// TIA Portal project "HEAT-1-CADIZ-V30" (V20) (continued)
VERSION : 0.1
// stored: InstanceOfName ToolChange
"ToolChange"
BEGIN
END_DATA_BLOCK

DATA_BLOCK "ToolChangeMarker_DB"   // DB40
{ S7_Optimized_Access := 'TRUE' }
VERSION : 0.1
// stored: InstanceOfName ToolChange
"ToolChange"
BEGIN
END_DATA_BLOCK

// folder: 30. Safety

DATA_BLOCK "InstMainSafety"   // DB1, F_DB
{ S7_Optimized_Access := 'TRUE' }
NAME : FUSI
VERSION : 0.1
// stored: InstanceOfName MainSafety
"MainSafety"
BEGIN
END_DATA_BLOCK

DATA_BLOCK "SafetyRobotDb"   // DB3, F_DB
{ S7_Optimized_Access := 'TRUE' }
VERSION : 0.1
BEGIN
END_DATA_BLOCK

DATA_BLOCK "EMERGENCIA_OPR_DB"   // DB41, F_DB
{ S7_Optimized_Access := 'TRUE' }
VERSION : 0.1
// stored: InstanceOfName EMERGENCIA_OPR
"EMERGENCIA_OPR"
BEGIN
END_DATA_BLOCK

DATA_BLOCK "EMERGENCIA_SETAS_DB"   // DB42, F_DB
{ S7_Optimized_Access := 'TRUE' }
VERSION : 0.1
// stored: InstanceOfName EMERGENCIA_SETAS
"EMERGENCIA_SETAS"
BEGIN
END_DATA_BLOCK

DATA_BLOCK "EMERGENCIAS_ANTENAS_DB"   // DB43, F_DB
{ S7_Optimized_Access := 'TRUE' }
VERSION : 0.1
// stored: InstanceOfName EMERGENCIAS_ANTENAS
"EMERGENCIAS_ANTENAS"
BEGIN
END_DATA_BLOCK

DATA_BLOCK "EMERGENCIA_GENERAL_DB"   // DB45, F_DB
{ S7_Optimized_Access := 'TRUE' }
VERSION : 0.1
// stored: InstanceOfName EMERGENCIA_GENERAL
"EMERGENCIA_GENERAL"
BEGIN
END_DATA_BLOCK

DATA_BLOCK "GESTION_BARRERAS_DB"   // DB46, F_DB
{ S7_Optimized_Access := 'TRUE' }
VERSION : 0.1
// stored: InstanceOfName GESTION_BARRERAS
"GESTION_BARRERAS"
BEGIN
END_DATA_BLOCK

// folder: 410. Festo cuba

DATA_BLOCK "HMI_CUBA_FESTO"   // DB12
{ S7_Optimized_Access := 'TRUE' }
VERSION : 0.1
   VAR
      HMI_Sensor_plato_giro_1 : Bool;
      HMI_Sensor_Plato_giro_2 : Bool;
      HMI_Sensor_plato_giro_3 : Bool;
      HMI_Sensor_ADN_bastidor_bloqueado_1 : Bool;
      HMI_Sensor_ADN_bastidor_desbloqueado_1 : Bool;
      HMI_Sensor_ADN_bastidor_bloqueado_2 : Bool;
      HMI_Sensor_ADN_bastidor_desbloqueado_2 : Bool;
      HMI_SENSOR_CRDSNU_BASTIDOR_BLOQUEADO_1 : Bool;
      HMI_SENSOR_CRDSNU_BASTIDOR_DESBLOQUEADO_1 : Bool;
      HMI_SENSOR_CRDSNU_BASTIDOR_BLOQUEADO_2 : Bool;
      HMI_SENSOR_CRDSNU_BASTIDOR_DESBLOQUEADO_2 : Bool;
      HMI_SENSOR_DSBG_BASTIDOR_ARRIBA_1 : Bool;
      HMI_SENSOR_DSBG_BASTIDOR_ABAJO_1 : Bool;
      HMI_SENSOR_DSBG_BASTIDOR_ARRIBA_2 : Bool;
      HMI_SENSOR_DSBG_BASTIDOR_ABAJO_2 : Bool;
      HMI_PULSADOR_SUBIR_1 : Bool;
      HMI_PULSADOR_BAJAR_1 : Bool;
      HMI_PULSADOR_SUBIR_2 : Bool;
      HMI_PULSADOR_BAJAR_2 : Bool;
      HMI_PULSADOR_BAJAR_3 : Bool;
      HMI_PULSADOR_BAJAR_4 : Bool;
      HMI_PULSADOR_BAJAR_5 : Bool;
      HMI_PULSADOR_BAJAR_6 : Bool;
      HMI_PULSADOR_BAJAR_7 : Bool;
      HMI_PULSADOR_BAJAR_8 : Bool;
      HMI_PULSADOR_BAJAR_9 : Bool;
      HMI_PULSADOR_BAJAR_10 : Bool;
      HMI_PULSADOR_BAJAR_11 : Bool;
      HMI_PULSADOR_BAJAR_12 : Bool;
      HMI_PULSADOR_BAJAR_13 : Bool;
      HMI_PULSADOR_BAJAR_14 : Bool;
      HMI_VALVULA_52_BIESTABLE_11 : Bool;
      HMI_VALVULA_52_BIESTABLE_12 : Bool;
      HMI_VALVULA_52_BIESTABLE_21 : Bool;
      HMI_VALVULA_52_BIESTABLE_22 : Bool;
      HMI_VÁLVULA_52_MONOESTABLE_1 : Bool;
      HMI_VÁLVULA_52_MONOESTABLE_2 : Bool;
      HMI_VÁLVULA_52_MONOESTABLE_3 : Bool;
      HMI_VÁLVULA_52_MONOESTABLE_4 : Bool;
      HMI_VÁLVULA_52_MONOESTABLE_5 : Bool;
      HMI_VÁLVULA_52_MONOESTABLE_6 : Bool;
      HMI_VÁLVULA_52_MONOESTABLE_7 : Bool;
      HMI_VÁLVULA_52_MONOESTABLE_8 : Bool;
      HMI_VÁLVULA_52_MONOESTABLE_9 : Bool;
      HMI_VÁLVULA_52_MONOESTABLE_10 : Bool;
      HMI_VÁLVULA_52_MONOESTABLE_11 : Bool;
      HMI_VÁLVULA_52_MONOESTABLE_12 : Bool;
      HMI_VÁLVULA_52_MONOESTABLE_13 : Bool;
      HMI_VÁLVULA_52_MONOESTABLE_14 : Bool;
      HMI_VÁLVULA_52_MONOESTABLE_15 : Bool;
      HMI_VÁLVULA_52_MONOESTABLE_16 : Bool;
      HMI_VÁLVULA_52_MONOESTABLE_17 : Bool;
      HMI_VÁLVULA_52_MONOESTABLE_18 : Bool;
      HMI_VÁLVULA_52_MONOESTABLE_19 : Bool;
      HMI_VÁLVULA_52_MONOESTABLE_20 : Bool;
      HMI_VÁLVULA_52_MONOESTABLE_21 : Bool;
      HMI_VÁLVULA_52_MONOESTABLE_22 : Bool;
      HMI_VÁLVULA_52_MONOESTABLE_23 : Bool;
      HMI_VÁLVULA_52_MONOESTABLE_24 : Bool;
      HMI_VÁLVULA_52_MONOESTABLE_25 : Bool;
      HMI_VÁLVULA_52_MONOESTABLE_26 : Bool;
      HMI_VÁLVULA_52_MONOESTABLE_27 : Bool;
      HMI_VÁLVULA_52_MONOESTABLE_28 : Bool;
      Estado_giro_pos_1 : Bool;
      Estado_giro_pos_2 : Bool;
      Estado_giro_pos_3 : Bool;
      Estado_giro_pos_4 : Bool;
      Estado_giro_neg_1 : Bool;
      Estado_giro_neg_2 : Bool;
      Estado_giro_neg_3 : Bool;
      Estado_giro_neg_4 : Bool;
      Estado_giro_neg_0 : Bool := true;
      Estado_giro_pos_0 : Bool := true;
      GIRO_AUTOMATICO_HABILITADO : Bool;
      Giro_negativo_auto : Bool;
      Giro_positivo_auto : Bool;
   END_VAR
BEGIN
END_DATA_BLOCK

// folder: Achim

DATA_BLOCK "Achim_testPepaFrk_DB"   // DB19
{ S7_Optimized_Access := 'TRUE' }
VERSION : 0.1
// stored: InstanceOfName Achim_testPepaFrk
"Achim_testPepaFrk"
BEGIN
END_DATA_BLOCK

// folder: Eliminar

DATA_BLOCK "DB_Supervisor"   // DB9
{ S7_Optimized_Access := 'TRUE' }
VERSION : 0.1
   VAR
      Common : Struct
         plc_ok : Bool;
         supervisor_ok : Bool;
         system_ok : Bool;
         safety_ok : Bool;
         air_ok : Bool;
         insp_water_ok : Bool;
         tank_water_ok : Bool;
         robot_ok : Bool;
         step_plc : Int;
         step_supervisor : Int;
         error : Bool;
         reset_req : Bool;
      END_STRUCT;
      Identification : Struct   // pag 2
         carriage_id_req : Bool;   // Sup->PLC
         new_carriage_id : Bool;   // PLC->Sup
         id_req : Bool;   // Sup->PLC
         id_running : Bool;   // PLC->Sup
         id_ok : Bool;   // PLC->Sup
         teach_req : Bool;   // Sup->PLC
         system_ok : Bool;   // PLC->Sup (parte de id_ok)
         pa_check_req : Bool;   // Sup->PLC
         tcg_req : Bool;   // Sup->PLC
      END_STRUCT;
      Teaching : Struct   // pag 3
         teach_ready : Bool;   // PLC->Sup
         teach_running : Bool;   // Sup->PLC
         teach_state : Bool;   // Sup->PLC
         jump_start_us : Bool;   // PLC->Sup
      END_STRUCT;
      StartUs : Struct   // pag 4
         start_us_ready : Bool;   // PLC->Sup
         start_us_running : Bool;   // Sup->PLC
         start_us_state : Bool;   // Sup->PLC
      END_STRUCT;
      PACheck : Struct   // pag 5
         pa_check_ready : Bool;   // PLC->Sup
         elem_running : Bool;   // Sup->PLC
         elem_state : Bool;   // Sup->PLC
         bal_running : Bool;   // Sup->PLC
         bal_state : Bool;   // Sup->PLC
      END_STRUCT;
      Gain : Struct
         gain_ready : Bool;
         gain_running : Bool;
         gain_state : Bool;
      END_STRUCT;
      TCG_Check : Struct
         tcg_ready : Bool;
         tcg_running : Bool;
         tcg_next_step : Bool;
         jump_acq_ref : Bool;
         jump_tcg_adj : Bool;
      END_STRUCT;
      TCG_Adjust : Struct
         tcg_ready : Bool;
         jump_ref_acq : Bool;
      END_STRUCT;
      RefScan_Acq : Struct
         scan_ref_ready : Bool;
         scan_ref_running : Bool;
      END_STRUCT;
      InspScan : Struct
         scan_insp_ready : Bool;
         scan_insp_running : Bool;
         scan_insp_state : Bool;
         jump_ref_insp : Bool;
      END_STRUCT;
      RefScan_Verif : Struct
         scan_ref_ready : Bool;
         scan_ref_running : Bool;
         jump_start : Bool;
      END_STRUCT;
      Marking : Struct
         mark_req : Bool;
         mark_running : Bool;
         mark_state : Bool;
         jump_start : Bool;
         point_coordinates : Struct
            x : Real;
            y : Real;
            z : Real;
            "a" : Real;
            "b" : Real;
            c : Real;
         END_STRUCT;
      END_STRUCT;
   END_VAR
BEGIN
END_DATA_BLOCK

// folder: System blocks/Program resources

DATA_BLOCK "IEC_Timer_0_DB"   // DB24
{ S7_Optimized_Access := 'TRUE' }
AUTHOR : Simatic
FAMILY : IEC
NAME : IEC_TMR
VERSION : 1.0
// stored: InstanceOfName IEC_TIMER
"IEC_TIMER"
BEGIN
END_DATA_BLOCK

DATA_BLOCK "IEC_Timer_0_DB_1"   // DB25
{ S7_Optimized_Access := 'TRUE' }
AUTHOR : Simatic
FAMILY : IEC
NAME : IEC_TMR
VERSION : 1.0
// stored: InstanceOfName IEC_TIMER
"IEC_TIMER"
BEGIN
END_DATA_BLOCK

DATA_BLOCK "IEC_Timer_0_DB_2"   // DB26
{ S7_Optimized_Access := 'TRUE' }
AUTHOR : Simatic
FAMILY : IEC
NAME : IEC_TMR
VERSION : 1.0
// stored: InstanceOfName IEC_TIMER
"IEC_TIMER"
BEGIN
END_DATA_BLOCK

DATA_BLOCK "IEC_Timer_0_DB_3"   // DB29
{ S7_Optimized_Access := 'TRUE' }
AUTHOR : Simatic
FAMILY : IEC
NAME : IEC_TMR
VERSION : 1.0
// stored: InstanceOfName IEC_TIMER
"IEC_TIMER"
BEGIN
END_DATA_BLOCK

DATA_BLOCK "IEC_Timer_0_DB_4"   // DB30
{ S7_Optimized_Access := 'TRUE' }
AUTHOR : Simatic
FAMILY : IEC
NAME : IEC_TMR
VERSION : 1.0
// stored: InstanceOfName IEC_TIMER
"IEC_TIMER"
BEGIN
END_DATA_BLOCK

DATA_BLOCK "IEC_Timer_0_DB_5"   // DB31
{ S7_Optimized_Access := 'TRUE' }
AUTHOR : Simatic
FAMILY : IEC
NAME : IEC_TMR
VERSION : 1.0
// stored: InstanceOfName IEC_TIMER
"IEC_TIMER"
BEGIN
END_DATA_BLOCK

DATA_BLOCK "IEC_Timer_0_DB_6"   // DB33
{ S7_Optimized_Access := 'TRUE' }
AUTHOR : Simatic
FAMILY : IEC
NAME : IEC_TMR
VERSION : 1.0
// stored: InstanceOfName IEC_TIMER
"IEC_TIMER"
BEGIN
END_DATA_BLOCK

DATA_BLOCK "IEC_Timer_0_DB_7"   // DB34
{ S7_Optimized_Access := 'TRUE' }
AUTHOR : Simatic
FAMILY : IEC
NAME : IEC_TMR
VERSION : 1.0
// stored: InstanceOfName IEC_TIMER
"IEC_TIMER"
BEGIN
END_DATA_BLOCK

DATA_BLOCK "IEC_Timer_0_DB_8"   // DB35
{ S7_Optimized_Access := 'TRUE' }
AUTHOR : Simatic
FAMILY : IEC
NAME : IEC_TMR
VERSION : 1.0
// stored: InstanceOfName IEC_TIMER
"IEC_TIMER"
BEGIN
END_DATA_BLOCK

DATA_BLOCK "IEC_Timer_0_DB_9"   // DB36
{ S7_Optimized_Access := 'TRUE' }
AUTHOR : Simatic
FAMILY : IEC
NAME : IEC_TMR
VERSION : 1.0
// stored: InstanceOfName IEC_TIMER
"IEC_TIMER"
BEGIN
END_DATA_BLOCK

DATA_BLOCK "IEC_Timer_0_DB_10"   // DB38
{ S7_Optimized_Access := 'TRUE' }
AUTHOR : Simatic
FAMILY : IEC
NAME : IEC_TMR
VERSION : 1.0
// stored: InstanceOfName IEC_TIMER
"IEC_TIMER"
BEGIN
END_DATA_BLOCK

// folder: (top level)

ORGANIZATION_BLOCK "Startup"   // OB100, LAD, Startup
TITLE = "Complete Restart"
{ S7_Optimized_Access := 'TRUE' }
VERSION : 0.1
   VAR_INPUT
      LostRetentive : Bool;   // True if retentive data are lost
      LostRTC : Bool;   // True if date and time are lost
   END_VAR
BEGIN

REGION Network 1 (SCL): // ====================== READ (%I) ======================
   // // —— Enlaza estos símbolos a tus %I en el árbol de dispositivos ——
   //   // EStop_DI, SafeDoor_DI, AirPressure_DI, WaterInsp_DI, WaterTank_DI, RobotReady_DI, ...
   "$MOVE_ENABLE" := TRUE;
END_REGION
END_ORGANIZATION_BLOCK

// folder: 10. System

FUNCTION_BLOCK "SeqManager"   // FB20, LAD
{ S7_Optimized_Access := 'TRUE' }
VERSION : 0.1
   VAR_INPUT
      systemArmed : Bool;
      autoBusy : Bool;
      servBusy : Bool;
      modeRequest : UInt;
      modeReqSeq : UInt;
   END_VAR
   VAR_OUTPUT
      modeEffective : UInt;
      startAutoExt : Bool;
      enterCellCase1 : Bool;
      enterCellCase2 : Bool;
   END_VAR
   VAR
      lastSeq : UInt;
      safeAllOk : Bool;
      acceptSrv : Bool;
      acceptAuto : Bool;
      firstScan : Bool := true;
   END_VAR
BEGIN

REGION Network 1 (SCL)
   // ----------------- 0) Inicialización por scan -----------------
   "PlcStatus".exec.accepted := FALSE; // pulso hacia la HMI
   "PlcStatus".exec.done := FALSE;    // pulso hacia la HMI

   // Clave: forzamos a FALSE por defecto para que al conceder se produzca pulso
   #startAutoExt := FALSE;
   #enterCellCase2 := FALSE;
   #enterCellCase1 := FALSE;

   // ----------------- 1) Inicialización primera pasada -----------------
   IF  #firstScan THEN
       #firstScan := FALSE;
       #lastSeq := #modeReqSeq;     // ignorar residuos SOLO al arrancar
   END_IF;

   #safeAllOk := #systemArmed;

   // Condición global de seguridad (quedar por ajustar)
   #safeAllOk := #systemArmed;


   IF #modeRequest = 3 THEN
       //#startAutoExt := TRUE;
       #lastSeq := #lastSeq + 1;
       // 5) Handshake a la HMI con el MISMO seq que se recibió
   END_IF;

   // ----------------- 2) Procesar SOLO peticiones nuevas (por secuencia) ----
   IF #modeReqSeq <> #lastSeq THEN
       #lastSeq := #modeReqSeq;

       CASE #modeRequest OF
           1: // ======= Conceder control a KukaControl =========
               // Requisito: que el otro lado (Supervisor) esté ocioso (Queda por ajustar)
               IF #safeAllOk AND (NOT #autoBusy) THEN

                   // 1) Fijar modo efectivo → AutoExtSeq cargará PGNO = 1
                   #modeEffective := USINT#1;

                   // 2) Aún no estamos listos hasta que AutoExtSeq termine
                   "PlcStatus".mode.ready := FALSE;

                   // 3) Señal PNIO al robot para que salga del bucle autoloop.src (CASE 1 del cell.src)
                   #enterCellCase1 := TRUE;

                   // 4) Arranque de AutoExt: PULSO 1-scan a %M770.0
                   #startAutoExt := TRUE;

                   // 5) Handshake a la HMI con el MISMO seq que se recibió
                   "PlcStatus".exec.ackSeq := #modeReqSeq;
                   "PlcStatus".exec.accepted := TRUE;  // 1 scan
                   "PlcStatus".exec.done := TRUE;  // 1 scan
               END_IF;

           2: // ======= Conceder control a Supervisor/VisualScan =========
               // Requisito: que KukaControl esté ocioso
               IF #safeAllOk AND (NOT #servBusy) THEN

                   // 1) Fijar modo efectivo → AutoExtSeq cargará PGNO = 2
                   #modeEffective := USINT#2;

                   // 2) Aún no estamos listos hasta que AutoExtSeq termine
                   "PlcStatus".mode.ready := FALSE;

                   // 3) Señal PNIO al robot para que salga del bucle actual autoloopsup.src (CASE 2 del cell.src)
                   #enterCellCase2 := TRUE;

                   // 4) Arranque de AutoExt: PULSO 1-scan a %M770.0
                   #startAutoExt := TRUE;

                   // 5) Handshake a la HMI
                   "PlcStatus".exec.ackSeq := #modeReqSeq;
                   "PlcStatus".exec.accepted := TRUE;
                   "PlcStatus".exec.done := TRUE;
               END_IF;
       END_CASE;

   END_IF;
END_REGION
END_FUNCTION_BLOCK

FUNCTION_BLOCK "KukaControlSeq"   // FB21, LAD
{ S7_Optimized_Access := 'TRUE' }
VERSION : 0.1
   VAR
      rEnterAuto : R_TRIG;
   END_VAR
   VAR_TEMP
      _clear990 : Bool;
   END_VAR
BEGIN

REGION Network 2: Envia posiciones a la aplicacion KukaControl
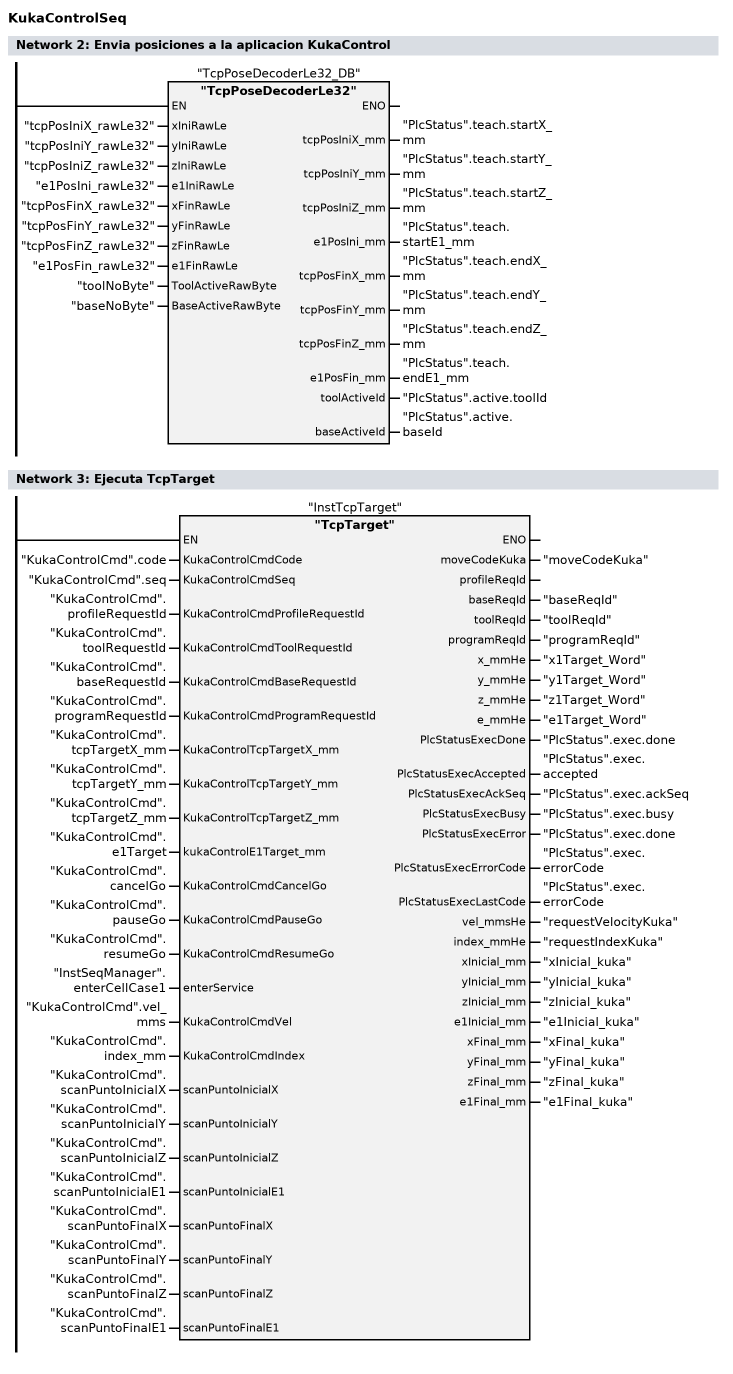
   RUNG wire#powerrail
      "TcpPoseDecoderLe32_DB"(xIniRawLe := "tcpPosIniX_rawLe32", yIniRawLe := "tcpPosIniY_rawLe32", zIniRawLe := "tcpPosIniZ_rawLe32", e1IniRawLe := "e1PosIni_rawLe32", xFinRawLe := "tcpPosFinX_rawLe32", yFinRawLe := "tcpPosFinY_rawLe32", zFinRawLe := "tcpPosFinZ_rawLe32", e1FinRawLe := "e1PosFin_rawLe32", ToolActiveRawByte := "toolNoByte", BaseActiveRawByte := "baseNoByte", tcpPosIniX_mm => "PlcStatus".teach.startX_mm, tcpPosIniY_mm => "PlcStatus".teach.startY_mm, tcpPosIniZ_mm => "PlcStatus".teach.startZ_mm, e1PosIni_mm => "PlcStatus".teach.startE1_mm, tcpPosFinX_mm => "PlcStatus".teach.endX_mm, tcpPosFinY_mm => "PlcStatus".teach.endY_mm, tcpPosFinZ_mm => "PlcStatus".teach.endZ_mm, e1PosFin_mm => "PlcStatus".teach.endE1_mm, toolActiveId => "PlcStatus".active.toolId, baseActiveId => "PlcStatus".active.baseId)
   END_RUNG
   // the same network as SCL:
   "TcpPoseDecoderLe32_DB"(xIniRawLe := "tcpPosIniX_rawLe32",   // "TcpPoseDecoderLe32"
                           yIniRawLe := "tcpPosIniY_rawLe32",
                           zIniRawLe := "tcpPosIniZ_rawLe32",
                           e1IniRawLe := "e1PosIni_rawLe32",
                           xFinRawLe := "tcpPosFinX_rawLe32",
                           yFinRawLe := "tcpPosFinY_rawLe32",
                           zFinRawLe := "tcpPosFinZ_rawLe32",
                           e1FinRawLe := "e1PosFin_rawLe32",
                           ToolActiveRawByte := "toolNoByte",
                           BaseActiveRawByte := "baseNoByte",
                           tcpPosIniX_mm => "PlcStatus".teach.startX_mm,
                           tcpPosIniY_mm => "PlcStatus".teach.startY_mm,
                           tcpPosIniZ_mm => "PlcStatus".teach.startZ_mm,
                           e1PosIni_mm => "PlcStatus".teach.startE1_mm,
                           tcpPosFinX_mm => "PlcStatus".teach.endX_mm,
                           tcpPosFinY_mm => "PlcStatus".teach.endY_mm,
                           tcpPosFinZ_mm => "PlcStatus".teach.endZ_mm,
                           e1PosFin_mm => "PlcStatus".teach.endE1_mm,
                           toolActiveId => "PlcStatus".active.toolId,
                           baseActiveId => "PlcStatus".active.baseId);
END_REGION

REGION Network 3: Ejecuta TcpTarget
   RUNG wire#powerrail
      "InstTcpTarget"(KukaControlCmdCode := "KukaControlCmd".code, KukaControlCmdSeq := "KukaControlCmd".seq, KukaControlCmdProfileRequestId := "KukaControlCmd".profileRequestId, KukaControlCmdToolRequestId := "KukaControlCmd".toolRequestId, KukaControlCmdBaseRequestId := "KukaControlCmd".baseRequestId, KukaControlCmdProgramRequestId := "KukaControlCmd".programRequestId, KukaControlTcpTargetX_mm := "KukaControlCmd".tcpTargetX_mm, KukaControlTcpTargetY_mm := "KukaControlCmd".tcpTargetY_mm, KukaControlTcpTargetZ_mm := "KukaControlCmd".tcpTargetZ_mm, kukaControlE1Target_mm := "KukaControlCmd".e1Target, KukaControlCmdCancelGo := "KukaControlCmd".cancelGo, KukaControlCmdPauseGo := "KukaControlCmd".pauseGo, KukaControlCmdResumeGo := "KukaControlCmd".resumeGo, enterService := "InstSeqManager".enterCellCase1, KukaControlCmdVel := "KukaControlCmd".vel_mms, KukaControlCmdIndex := "KukaControlCmd".index_mm, scanPuntoInicialX := "KukaControlCmd".scanPuntoInicialX, scanPuntoInicialY := "KukaControlCmd".scanPuntoInicialY, scanPuntoInicialZ := "KukaControlCmd".scanPuntoInicialZ, scanPuntoInicialE1 := "KukaControlCmd".scanPuntoInicialE1, scanPuntoFinalX := "KukaControlCmd".scanPuntoFinalX, scanPuntoFinalY := "KukaControlCmd".scanPuntoFinalY, scanPuntoFinalZ := "KukaControlCmd".scanPuntoFinalZ, scanPuntoFinalE1 := "KukaControlCmd".scanPuntoFinalE1, moveCodeKuka => "moveCodeKuka", profileReqId =>, baseReqId => "baseReqId", toolReqId => "toolReqId", programReqId => "programReqId", x_mmHe => "x1Target_Word", y_mmHe => "y1Target_Word", z_mmHe => "z1Target_Word", e_mmHe => "e1Target_Word", PlcStatusExecDone => "PlcStatus".exec.done, PlcStatusExecAccepted => "PlcStatus".exec.accepted, PlcStatusExecAckSeq => "PlcStatus".exec.ackSeq, PlcStatusExecBusy => "PlcStatus".exec.busy, PlcStatusExecError => "PlcStatus".exec.done, PlcStatusExecErrorCode => "PlcStatus".exec.errorCode, PlcStatusExecLastCode => "PlcStatus".exec.errorCode, vel_mmsHe => "requestVelocityKuka", index_mmHe => "requestIndexKuka", xInicial_mm => "xInicial_kuka", yInicial_mm => "yInicial_kuka", zInicial_mm => "zInicial_kuka", e1Inicial_mm => "e1Inicial_kuka", xFinal_mm => "xFinal_kuka", yFinal_mm => "yFinal_kuka", zFinal_mm => "zFinal_kuka", e1Final_mm => "e1Final_kuka")
   END_RUNG
   // the same network as SCL:
   "InstTcpTarget"(KukaControlCmdCode := "KukaControlCmd".code,   // "TcpTarget"
                   KukaControlCmdSeq := "KukaControlCmd".seq,
                   KukaControlCmdProfileRequestId := "KukaControlCmd".profileRequestId,
                   KukaControlCmdToolRequestId := "KukaControlCmd".toolRequestId,
                   KukaControlCmdBaseRequestId := "KukaControlCmd".baseRequestId,
                   KukaControlCmdProgramRequestId := "KukaControlCmd".programRequestId,
                   KukaControlTcpTargetX_mm := "KukaControlCmd".tcpTargetX_mm,
                   KukaControlTcpTargetY_mm := "KukaControlCmd".tcpTargetY_mm,
                   KukaControlTcpTargetZ_mm := "KukaControlCmd".tcpTargetZ_mm,
                   kukaControlE1Target_mm := "KukaControlCmd".e1Target,
                   KukaControlCmdCancelGo := "KukaControlCmd".cancelGo,
                   KukaControlCmdPauseGo := "KukaControlCmd".pauseGo,
                   KukaControlCmdResumeGo := "KukaControlCmd".resumeGo,
                   enterService := "InstSeqManager".enterCellCase1,
                   KukaControlCmdVel := "KukaControlCmd".vel_mms,
                   KukaControlCmdIndex := "KukaControlCmd".index_mm,
                   scanPuntoInicialX := "KukaControlCmd".scanPuntoInicialX,
                   scanPuntoInicialY := "KukaControlCmd".scanPuntoInicialY,
                   scanPuntoInicialZ := "KukaControlCmd".scanPuntoInicialZ,
                   scanPuntoInicialE1 := "KukaControlCmd".scanPuntoInicialE1,
                   scanPuntoFinalX := "KukaControlCmd".scanPuntoFinalX,
                   scanPuntoFinalY := "KukaControlCmd".scanPuntoFinalY,
                   scanPuntoFinalZ := "KukaControlCmd".scanPuntoFinalZ,
                   scanPuntoFinalE1 := "KukaControlCmd".scanPuntoFinalE1,
                   moveCodeKuka => "moveCodeKuka",
                   baseReqId => "baseReqId",
                   toolReqId => "toolReqId",
                   programReqId => "programReqId",
                   x_mmHe => "x1Target_Word",
                   y_mmHe => "y1Target_Word",
                   z_mmHe => "z1Target_Word",
                   e_mmHe => "e1Target_Word",
                   PlcStatusExecDone => "PlcStatus".exec.done,
                   PlcStatusExecAccepted => "PlcStatus".exec.accepted,
                   PlcStatusExecAckSeq => "PlcStatus".exec.ackSeq,
                   PlcStatusExecBusy => "PlcStatus".exec.busy,
                   PlcStatusExecError => "PlcStatus".exec.done,
                   PlcStatusExecErrorCode => "PlcStatus".exec.errorCode,
                   PlcStatusExecLastCode => "PlcStatus".exec.errorCode,
                   vel_mmsHe => "requestVelocityKuka",
                   index_mmHe => "requestIndexKuka",
                   xInicial_mm => "xInicial_kuka",
                   yInicial_mm => "yInicial_kuka",
                   zInicial_mm => "zInicial_kuka",
                   e1Inicial_mm => "e1Inicial_kuka",
                   xFinal_mm => "xFinal_kuka",
                   yFinal_mm => "yFinal_kuka",
                   zFinal_mm => "zFinal_kuka",
                   e1Final_mm => "e1Final_kuka");
END_REGION

REGION Network 4 (SCL)
   IF #_clear990 THEN
       "KukaControlCmd".code := 0;                     // no “ensucia” el DB
       #_clear990 := FALSE;
   END_IF;
END_REGION
END_FUNCTION_BLOCK

FUNCTION_BLOCK "SupervisorSeq"   // FB22, LAD
{ S7_Optimized_Access := 'TRUE' }
VERSION : 0.1
   VAR_INPUT
      T_Heartbeat : Time := T#1000ms;   // Periodo del heartbeat PLC
      T_IdCheck : Time := T#2000ms;   // Duración simulada de Identification (comprobaciones)
      QR_Ready : Bool := true;   // Hay un ID de carrito leído
      CarriageID : String := 'null';   // ID de carrito leído por QR
      SupervisorCmdReqCarriageId : Bool;
      SupervisorCmdReqId : Bool;
      SupervisorCmdPns : String;
      SupervisorCmdReferencePart : String;
      SupervisorCmdEndEffector : Int;
      SupervisorCmdUtTech : UInt;
      SupervisorCmdTeachReq : Bool;
      SupervisorCmdPaCheckReq : Bool;
      SupervisorCmdTcgReq : Bool;
      SupervisorCmdStartUsRunning : Bool;
      SupervisorCmdStateUs : Bool;
      SupervisorCmdGainRunning : Bool;
      SupervisorCmdGainState : Bool;
      TeachAtStart : Bool;   // Teaching (pág. 4): robot en punto de inicio de la siguiente trayectoria
      kukaAtPerspexPos : Bool;   // PA check (Perspex) y Balancing (pág. 6): Robot posicionado en Perspex
      kukaAtGainPos : Bool;   // Gain (pág. 7) -Robot posicionado para Gain
      kukaAtTCGPos : Bool;   // TCG (pág. 8) — multiposición Robot en la posición TCG actual
      kukaAtRefScanStartPos : Bool;   // Robot listo para Scan Ref
      kukaAtInspScanStartPos : Bool;   // Robot listo para Scan Insp
      kukaRefScanFinished : Bool;   // Trayectoria de referencia terminada (robot/UT)
      kukaInspScanFinished : Bool;   // Trayectoria de inspección terminada (robot/UT)
      StartUSReady : Bool := TRUE;   // StartUS (pág. 5): end-effector y precondiciones listas -- True cuando “previous task done”
      MarkingDone : Bool;   // Pre-eval / marcado (pág. 13) -Resultado del marcado (true=OK)
      CmdStopUS : Bool;   // Orden local para Stop US
      CmdBreakUS : Bool;   // Pulso local Break US
      CmdUnbreakUS : Bool;   // Pulso local Unbreak US
   END_VAR
   VAR_OUTPUT
      ActiveStep : Int;   // Espejo local de PLC.step_plc
      PlcStatusStepPlc : Int;
      PlcStatusCarriageId : String;
      PlcStatusNewCarriageId : Bool;
      PlcStatusIdRunning : Bool;
      PlcStatusIdOk : Bool;
      PlcStatusStartUsReady : Bool;
      PlcStatusGainReady : Bool;
      moveCodeKuka : Word;
      toolReqId : Int;
      programReqId : Word;
      AckSourceDbg : Int;   // Código de fuente de ACK (debug local)
      TCG_NextPosReq : Bool;   // PULSO 1 ciclo: mover a la SIGUIENTE posición TCG
      TCG_AdjustMode : Bool;   // LATCH: TRUE mientras estamos en “ajuste TCG”
   END_VAR
   VAR
      tHeartbeat : TON_TIME;
      hbGate : Bool;
      prevStep : Int := -32768;
      firstScan : Bool;
      teachWasRunning : Bool;
      startUSWasRunning : Bool;
      scanRefWasRunning : Bool;
      scanInspWasRunning : Bool;
      L_IdEvalDone : Bool;   // // Identification: ya evalué reqId
      carriageLatched : Bool;
      validScanParams : Bool;
      waitingNextTCGPos : Bool;
      Cfg_Pns : String;
      Cfg_ReferencePart : String;
      Cfg_EndEffector : Int;
      Cfg_UtTeach : UInt;
      Cfg_TeachReq : Bool;
      Cfg_PaCheckReq : Bool;
      Cfg_TcgReq : Bool;
      PartProgIdx : UInt := 1;   // // index de programa INSP (pieza)
      RefProgIdx : UInt := 1;   // // index de programa REF (pieza)
      tcgIndex : UInt := 1;   // // posición TCG actual
      WantCode_uint : UInt;
      WantProgRequestId : Int;
      WantToolRequestId : Int;
      WantIndex : UInt;
      state : Int;
      lastSeq : UInt;
      SupervisorCmdSeq : UInt;
      handshakeStep : Int;   // // Handshake Manager (Gestión de Acknowledge 4-vías y sincronización)
      paBalSubStep : Int;   // // Sub-estados para pasos complejos
      gainSubStep : Int;
      markingSubStep : Int;
      tempNextStep : Int;   // // Almacena el siguiente paso principal
   END_VAR
   VAR_TEMP
      _clear990 : Bool;
      code_int : UInt;
   END_VAR
   VAR CONSTANT
      cSTEP_ID : Int := 1;   // // Pasos (según resumen del PDF, pág. 1)
      cSTEP_TEACH : Int := 2;
      cSTEP_STARTUS : Int := 3;
      cSTEP_PA_BAL : Int := 4;
      cSTEP_GAIN : Int := 5;
      cSTEP_TCG : Int := 6;
      cSTEP_SCAN_REF : Int := 7;
      cSTEP_SCAN_INSP : Int := 8;
      cSTEP_SCAN_REF_VERIF : Int := 9;
      cSTEP_PRE_EVAL : Int := 10;
      cKUKA_REQ_TOOL : UInt := 201;
      cKUKA_GOTO_PERSPEX : UInt := 412;   // mover a Perspex (usa punto enseñado en KRC)
      cKUKA_GOTO_GAIN : UInt := 413;   // mover a Gain
      cKUKA_GOTO_TCG : UInt := 414;   // mover a posición TCG (ARG = index)
      cKUKA_GOTO_REF_START : UInt := 420;   // mover a inicio de Ref (ARG = RefProgIdx)
      cKUKA_GOTO_INSP_START : UInt := 421;   // mover a inicio de Insp (ARG = PartProgIdx)
      cKUKA_RUN_REF_PATH : UInt := 432;   // ejecutar trayectoria de Ref (ARG = RefProgIdx)
      cKUKA_RUN_INSP_PATH : UInt := 433;   // ejecutar trayectoria de Insp (ARG = PartProgIdx)
      cKUKA_GOTO_SAF : UInt := 100;
      cKUKA_RETRACT_PERSPEX : UInt := 101;
      cKUKA_RETRACT_GAIN : UInt := 102;
      cKUKA_RETRACT_TCG : UInt := 103;
      cKUKA_MARK_POINT : UInt := 501;
      cTOOL_MARKER : Int := 3;
   END_VAR
BEGIN

REGION Network 1 (SCL)
   // ------------------------------------------------------------------
   // 0) Servicios globales (Heartbeat, housekeeping) — vars generales (pág. 2)
   // ------------------------------------------------------------------

   // Heartbeat PLC: toggle con TON (patrón de "compuerta")
   // hbGate se pone TRUE -> TON corre hasta PT -> tHeartbeat.Q = TRUE -> togglamos
   // y bajamos hbGate para reiniciar el ciclo.
   #tHeartbeat(IN := #hbGate,
               PT := #T_Heartbeat);
   IF NOT #hbGate THEN
       #hbGate := TRUE;
   ELSIF #tHeartbeat.Q THEN
       "PlcStatus".heartbeatPlc := NOT "PlcStatus".heartbeatPlc;
       #hbGate := FALSE;
   END_IF;

   // Normalizar paso y espejarlo a salida
   IF (#PlcStatusStepPlc < #cSTEP_ID) OR (#PlcStatusStepPlc > #cSTEP_PRE_EVAL) THEN
       #PlcStatusStepPlc := #cSTEP_ID;
   END_IF;
   #ActiveStep := #PlcStatusStepPlc;

   // firstScan: 1 ciclo al entrar en cada paso -> útil para resets seguros
   #firstScan := (#PlcStatusStepPlc <> #prevStep);
   IF #firstScan THEN
       // Limpiamos cualquier "ready/start" que no deba arrastrarse al paso nuevo
       "PlcStatus".startUsReady := FALSE;
       "PlcStatus".stopUsReady := FALSE;
       "PlcStatus".paCheckReady := FALSE;
       "PlcStatus".gainReady := FALSE;
       "PlcStatus".tcgReady := FALSE;
       "PlcStatus".scanRefStart := FALSE;
       "PlcStatus".scanInspStart := FALSE;
       "PlcStatus".markRunning := FALSE;
       "PlcStatus".acknowledge := FALSE; // [MEJORA] Reset Acknowledge

       // Latches de “estaba corriendo”  (Solo los necesarios)
       #teachWasRunning := FALSE;
       #startUSWasRunning := FALSE;
       #scanRefWasRunning := FALSE;
       #scanInspWasRunning := FALSE;

       // [MEJORA] Reset de Sub-estados y Handshake Manager
       #paBalSubStep := 0;
       #gainSubStep := 0;
       #markingSubStep := 0;
       #handshakeStep := 0;


       // Identification
       "PlcStatus".idRunning := FALSE;
       #L_IdEvalDone := FALSE;

       // TCG
       // 
       #waitingNextTCGPos := FALSE; // Ya no se usa, reemplazado por tcgSubStep
       IF "PlcStatus".stepPlc <> #cSTEP_TCG THEN
           #tcgIndex := 1;
       END_IF;

       // Vaciar slot de orden pendiente a robot
       #WantCode_uint := 0;
       #WantProgRequestId := 0;
       #WantToolRequestId := 0;
       #WantIndex := 0;

       #prevStep := #PlcStatusStepPlc;
   END_IF;

   // ------------------------------------------------------------------
   //[1] MÁQUINA DE ESTADOS (OPC UA + disparos al KUKA por goTrigger)
   // ------------------------------------------------------------------
   CASE #PlcStatusStepPlc OF

           // ===============================================================
           // 1) IDENTIFICATION (pág. 3)
           // ===============================================================
           // ---------- Handshake de carriageID //-----------
           // FÍSICO: lectura real de QR/PNs/params en KukaControl.
           // El PLC refleja ID leído y valida condiciones base (safety, agua, robot OK).
           // 1)Si Supervisor.req_carriage_id = TRUE -> el PLC debe mandar:
           //   PLC.carriage_Id (string) y levanta PLC.new_carriage_Id = TRUE mientras dure la petición
           // 2) Al bajar la petición (Supervisor.req_carriage_id = FALSE) , el PLC
           // baja new_carriage_Id y deja de enviar.

       #cSTEP_ID:

           //1)si Supervisor.req_carriage_id=TRUE, el PLC publica PLC.carriage_Id y levanta PLC.new_carriage_Id
           IF #SupervisorCmdReqCarriageId THEN
               IF #QR_Ready AND NOT #carriageLatched  THEN
                   #CarriageID := 'SPUL-MP-01029-000-UTEN';
                   #PlcStatusCarriageId := #CarriageID; // escribimos el ID leído
                   #PlcStatusNewCarriageId := TRUE;     // “ID listo”
                   #carriageLatched  := TRUE;              // evita rearmar en el mismo pulso
               END_IF;
           ELSE
               // fin del handshake
               #PlcStatusNewCarriageId := FALSE;
               #carriageLatched  := FALSE;
           END_IF;


           //----------- Handshake de req_id -----------
           // 3)cuando Supervisor.req_id sube por primera vez, tu FB congela receta:
           // 4) Resuelve índices de programa por pieza (tu mapeo PIEZA1/2/3)
           // 5)Cuando req_id baja:
           //  5.1)Calcula PLC.id_ok con enclavamientos/servicios/robot OK y rango válido de herramienta
           //  5.2)Decide
           //      id_ok=FALSE → se queda en Identification (ciclo cancelado).
           //      id_ok=TRUE & teach_req=TRUE → iría a Teaching.
           //      id_ok=TRUE & teach_req=FALSE → StartUS.

           // Espejo de “en curso”: mientras req_id = TRUE, id_running = TRUE
           IF #SupervisorCmdReqId THEN
               #PlcStatusIdRunning := TRUE;
           END_IF;

